(* Logix 5000 project; controller FV vendor 1 type 14 code 217 rev 31.11; software revision 31.00; part 56 of 63 *)
(* tags used below, declared in another part *)
   CWD : CHECKWORD_FLAGS;
   FV_B42 : INT[255];   // YSVCIP_FLG
   FV_B82 : INT[255];   // YSTFILL FL YST filling process flags
   FV_B82_0_2_OutputBit : BOOL;
   FV_B86 : INT[255];   // YSTCIP FL YST CIP process flag s
   FV_F8 : REAL[256];
   FV_N12 : INT[255];   // SYS_PARMS System Parameter Fil e
   FV_N136 : INT[50];   // YSV1, CURRENT FV DATA
   FV_N137 : INT[50];   // YSV2, CURRENT FV DATA
   FV_N138 : INT[50];   // YSV3, CURRENT FV DATA
   FV_N139 : INT[255];   // YST1
   FV_N140 : INT[255];   // YST2
   FV_N141 : INT[255];   // YSV1 DATA
   FV_N142 : INT[255];   // YSV2 DATA
   FV_N143 : INT[255];   // YSV3 DATA
   FV_N144 : INT[255];   // YST1 DATA
   FV_N145 : INT[255];   // YST2 DATA
   FV_N80 : INT[255];   // YSTFILL<PC YST filling data fro m PC
   FV_N81 : INT[255];   // YSTFILL>PC YST filling process data to PC and contr ol regs.
   FV_N88 : INT[255];   // YSP COMMS Data transferred to/ from yeast press PLC
   FV_R2V1 : PlantItem;   // R2V1
   FV_R2V2 : PlantItem;   // R2V2
   FV_T4 : TIMER[10];
   FV_WYT1R : PlantItem;   // WYT1R
   FV_WYT2R : PlantItem;   // WYT2R
   FV_WYTR1 : PlantItem;   // WYTR1
   FV_WYTR2 : PlantItem;   // WYTR2
   FV_YST01_LTX501_Fill_Lvl_OK : TIMER;
   FV_YST02_LTX501_Fill_Lvl_OK : TIMER;
   FV_YST1_HL_SP : DINT;
   FV_YST2_HL_SP : DINT;
   FV_YSV1CV : PlantItem;   // YSV1CV
   FV_YSV1R : PlantItem;   // YSV1R
   FV_YSV2CV : PlantItem;   // YSV2CV
   FV_YSV2R : PlantItem;   // YSV2R
   FV_YSV3R : PlantItem;   // YSV3R
   MV_YST_Levels : REAL[2];
   YST_BL_PMP_ON : BOOL;   // Blunger Pump
   YST_Confirm_Vent_connected : BOOL;
   YST_Vent_Connection_Confirmed : BOOL;
(* FV_Common, continued *)

   34: OTU(FV_B82[0].0);
   35: EQU(FV_N80[1],1)EQU(FV_N144[0],1)MOV(5,FV_N144[0]);
   36: EQU(FV_N80[1],2)EQU(FV_N145[0],1)MOV(5,FV_N145[0]);
   // Set current YSTs operation to storage
   37: JSR(FV_Set_FV_Datafile_Value,3,5,FV_N81[15],0);
   // Switch current YST's rouser mode to automatic
   38: JSR(FV_Set_FV_Datafile_Value,3,0,FV_N81[15],3);
   39: [CLR(FV_N81[16]) ,CLR(FV_N80[0]) ];
   40: MCR();
   // Copy current step to PC display register
   41: XIC(FV_B82[0].1)MOV(FV_N81[1],FV_N81[9]);
END_ROUTINE

ROUTINE FV_YSTFILL_MC_80   (* ladder *)
   // YST Filling Master Control Program YST filling command processor
   0: JSR(FV_YSTFILL_CP_81,0);
   // YST filling process control program
   1: XIC(FV_B82[0].0)JSR(FV_YSTFILL_PR_82,0);
   // Postscan filling process program
   2: XIO(FV_B82[0].0)OSR(FV_B82[0].2,FV_B82_0_2_OutputBit)XIC(FV_B82_0_2_OutputBit)[JSR(FV_YSTFILL_PR_82,0) ,MOV(99,FV_N88[1]) ];
END_ROUTINE

ROUTINE FV_YSTFILL_PR_82   (* ladder *)
   // YST Filling Process Control Program Step 10: Initialise
   0: XIC(FV_B82[0].1)EQU(FV_N81[1],10)MCR();
   1: [OTE(YST_Confirm_Vent_connected) ,XIC(YST_Vent_Connection_Confirmed) MOV(11,FV_N81[1]) ];
   2: MCR();
   // YST Filling Process Control Program Step 10: Initialise
   3: XIC(FV_B82[0].1)EQU(FV_N81[1],11)MCR();
   4: OTU(YST_Vent_Connection_Confirmed);
   5: MOV(10,FV_N81[3]);
   // Initialise pointer to current YST's data and attemperation files
   6: [ADD(FV_N80[1],143,FV_N81[15]) ,ADD(FV_N80[1],138,FV_N81[14]) ];
   // Set current YST's dirty flag
   7: JSR(FV_Set_Flag_In_FV_Datafile,3,FV_N81[15],1,0);
   8: MOV(20,FV_N81[1]);
   9: MCR();
   // Step 20: fill YST
   10: XIC(FV_B82[0].1)EQU(FV_N81[1],20)MCR();
   11: MOV(20,FV_N81[3]);
   // Drive Valves (Rung 8)
   12: [EQU(FV_N80[1],1) LEQ(MV_YST_Levels[0],FV_YST1_HL_SP) [TON(FV_YST01_LTX501_Fill_Lvl_OK,?,?) ,XIC(FV_YST01_LTX501_Fill_Lvl_OK.DN) [OTE(FV_WYTR1.DriveBits.0) ,XIO(FV_B86[0].1) OTE(FV_R2V1.DriveBits.1) ,XIC(FV_WYTR1.CW.[CWD.OPENFB]) OTL(YST_BL_PMP_ON) ] ] ,EQU(FV_N80[1],2) LEQ(MV_YST_Levels[1],FV_YST2_HL_SP) [TON(FV_YST02_LTX501_Fill_Lvl_OK,?,?) ,XIC(FV_YST02_LTX501_Fill_Lvl_OK.DN) [OTE(FV_WYTR2.DriveBits.0) ,XIO(FV_B86[0].1) OTE(FV_R2V2.DriveBits.1) ,XIC(FV_WYTR2.CW.[CWD.OPENFB]) OTL(YST_BL_PMP_ON) ] ] ];
   13: [OTE(FV_N81[2].5) ,XIC(FV_N80[0].5) MOV(30,FV_N81[1]) ];
   14: MCR();
   // Step 30: reset YST
   15: XIC(FV_B82[0].1)EQU(FV_N81[1],30)MCR();
   16: [JSR(FV_Set_FV_Datafile_Value,3,0,FV_N81[15],3) ,JSR(FV_Set_FV_Datafile_Value,3,5,FV_N81[15],0) ,CLR(FV_N81[16]) ,OTU(FV_N80[0].5) ,OTU(YST_BL_PMP_ON) ];
   17: MCR();
   // Check for alarms while running
   18: XIC(FV_B82[0].1)MCR();
   // High Level Alarm (Rung 15)
   19: [EQU(FV_N80[1],1) GEQ(MV_YST_Levels[0],FV_YST1_HL_SP) ,EQU(FV_N80[1],2) GEQ(MV_YST_Levels[1],FV_YST2_HL_SP) ][MOV(800,FV_N81[4]) ,MOV(FV_N80[1],FV_N81[5]) ];
   20: XIC(FV_N88[20].0)XIO(FV_N88[20].0)MOV(801,FV_N81[4]);
   21: [EQU(FV_N80[1],1) [XIC(FV_WYTR1.CW.[CWD.FAULT]) ,XIC(FV_R2V1.CW.[CWD.FAULT]) ] ,EQU(FV_N80[1],2) [XIC(FV_WYTR2.CW.[CWD.FAULT]) ,XIC(FV_R2V2.CW.[CWD.FAULT]) ] ,GRT(FV_N81[4],0) ][OTU(FV_B82[0].1) ,OTU(YST_BL_PMP_ON) ];
   22: XIC(FV_B82[0].1)MOV(FV_N80[1],FV_N88[1]);
   23: XIO(FV_B82[0].1)[MOV(4,FV_N81[0]) ,OTU(FV_N81[2].2) ,OTL(FV_N81[2].3) ,OTL(FV_N81[2].4) ,MOV(0,FV_N81[1]) ,MOV(99,FV_N88[1]) ,OTU(YST_BL_PMP_ON) ,OTU(YST_Vent_Connection_Confirmed) ];
   24: MCR();
END_ROUTINE

ROUTINE FV_YSV_ROUSE_112   (* ladder *)
   // ROUSING TIMERS Load Rouser On Period during storage from settings file
   0: MUL(FV_N12[6],1000,FV_T4[3].PRE);
   // Load Rouser Off Period during storage from settings file
   1: MUL(FV_N12[7],1000,FV_T4[4].PRE);
   // Enforce some minimum values on these timers
   2: LES(FV_T4[3].PRE,300000)MUL(300,1000,FV_T4[3].PRE);
   // Enforce some minimum values on these timers
   3: LES(FV_T4[4].PRE,300000)MUL(300,1000,FV_T4[4].PRE);
   // Cyclic timers for YSV rousing during storage
   4: XIO(FV_T4[4].DN)TON(FV_T4[3],?,?);
   5: XIC(FV_T4[3].DN)TON(FV_T4[4],?,?);
   // Load Rouser On Period during CIP from settings file
   6: MUL(FV_N12[8],1000,FV_T4[5].PRE);
   // Enforce some minimum values on these timers
   7: LES(FV_T4[5].PRE,600000)MUL(600,1000,FV_T4[5].PRE);
   // Rousing timer for CIP
   8: XIC(FV_B42[0].1)TON(FV_T4[5],?,?);
   // YSV 1 ROUSING Request rouser whilst attemporation active on this vesssel
   9: EQU(FV_N141[3],0)EQU(FV_N136[24],10)[[GRT(FV_N136[25],60) ,XIC(FV_YSV1R.DriveBits.0) GRT(FV_N136[25],45) ] ,LEQ(FV_N136[25],60) XIC(FV_T4[3].TT) ]OTE(FV_YSV1R.DriveBits.0);
   // Request rouser during CIP of this vessel
   10: EQU(FV_N141[3],0)EQU(FV_N141[0],3)XIC(FV_T4[5].TT)OTE(FV_YSV1R.DriveBits.1);
   // Request rouser if set to manual / continuous rouse
   11: EQU(FV_N141[3],1)OTE(FV_YSV1R.DriveBits.2);
   // YSV 2 ROUSING Request rouser whilst attemporation active on this vesssel
   12: EQU(FV_N142[3],0)EQU(FV_N137[24],10)[[GRT(FV_N137[25],60) ,XIC(FV_YSV2R.DriveBits.0) GRT(FV_N137[25],45) ] ,LEQ(FV_N137[25],60) XIC(FV_T4[3].TT) ]OTE(FV_YSV2R.DriveBits.0);
   // Request rouser during CIP of this vessel
   13: EQU(FV_N142[3],0)EQU(FV_N142[0],3)XIC(FV_T4[5].TT)OTE(FV_YSV2R.DriveBits.1);
   // Request rouser if set to manual / continuous rouse
   14: EQU(FV_N142[3],1)OTE(FV_YSV2R.DriveBits.2);
   // YSV 3 ROUSING Request rouser whilst attemporation active on this vesssel
   15: EQU(FV_N143[3],0)EQU(FV_N138[24],10)[[GRT(FV_N138[25],60) ,XIC(FV_YSV3R.DriveBits.0) GRT(FV_N138[25],45) ] ,LEQ(FV_N138[25],60) XIC(FV_T4[3].TT) ]OTE(FV_YSV3R.DriveBits.0);
   // Request rouser during CIP of this vessel
   16: EQU(FV_N143[3],0)EQU(FV_N143[0],3)XIC(FV_T4[5].TT)OTE(FV_YSV3R.DriveBits.1);
   // Request rouser if set to manual / continuous rouse
   17: EQU(FV_N143[3],1)OTE(FV_YSV3R.DriveBits.2);
   // YSTs 1 and 2 Rouser Control Request YST1 rouser if YST1 chilling active
   18: EQU(FV_N144[3],0)XIC(FV_N139[30].0)XIC(FV_YSV1CV.CW.[CWD.OUTPUT])OTE(FV_WYT1R.DriveBits.0);
   19: EQU(FV_N144[3],1)OTE(FV_WYT1R.DriveBits.1);
   // Request YST2 rouser if YST2 chilling active
   20: EQU(FV_N145[3],0)XIC(FV_N140[30].0)XIC(FV_YSV2CV.CW.[CWD.OUTPUT])OTE(FV_WYT2R.DriveBits.0);
   // Request YST2 rouser if rouser mode = manual on
   21: EQU(FV_N145[3],1)OTE(FV_WYT2R.DriveBits.1);
END_ROUTINE

ROUTINE FV_YSV_VOLUME_113   (* ladder *)
   // YSV 1
   0: EQU(FV_N141[7],0)MOV(10000,FV_N141[7]);
   1: MUL(FV_N141[7],0.1,FV_F8[3]);
   2: DIV(FV_N141[2],FV_F8[3],FV_F8[4]);
   3: MUL(FV_F8[4],1000.0,FV_F8[4]);
   4: GRT(FV_F8[4],32767.0)MOV(32767.0,FV_F8[4]);
   5: LES(FV_F8[4],0.0)MOV(0.0,FV_F8[4]);
   6: MOV(FV_F8[4],FV_N141[5]);
   // YSV 2
   7: EQU(FV_N142[7],0)MOV(10000,FV_N142[7]);
   8: MUL(FV_N142[7],0.1,FV_F8[3]);
   9: DIV(FV_N142[2],FV_F8[3],FV_F8[4]);
   10: MUL(FV_F8[4],1000.0,FV_F8[4]);
   11: GRT(FV_F8[4],32767.0)MOV(32767.0,FV_F8[4]);
   12: LES(FV_F8[4],0.0)MOV(0.0,FV_F8[4]);
   13: MOV(FV_F8[4],FV_N142[5]);
   // YSV 3
   14: EQU(FV_N143[7],0)MOV(10000,FV_N143[7]);
   15: MUL(FV_N143[7],0.1,FV_F8[3]);
   16: DIV(FV_N143[2],FV_F8[3],FV_F8[4]);
   17: MUL(FV_F8[4],1000.0,FV_F8[4]);
   18: GRT(FV_F8[4],32767.0)MOV(32767.0,FV_F8[4]);
   19: LES(FV_F8[4],0.0)MOV(0.0,FV_F8[4]);
   20: MOV(FV_F8[4],FV_N143[5]);
END_ROUTINE
